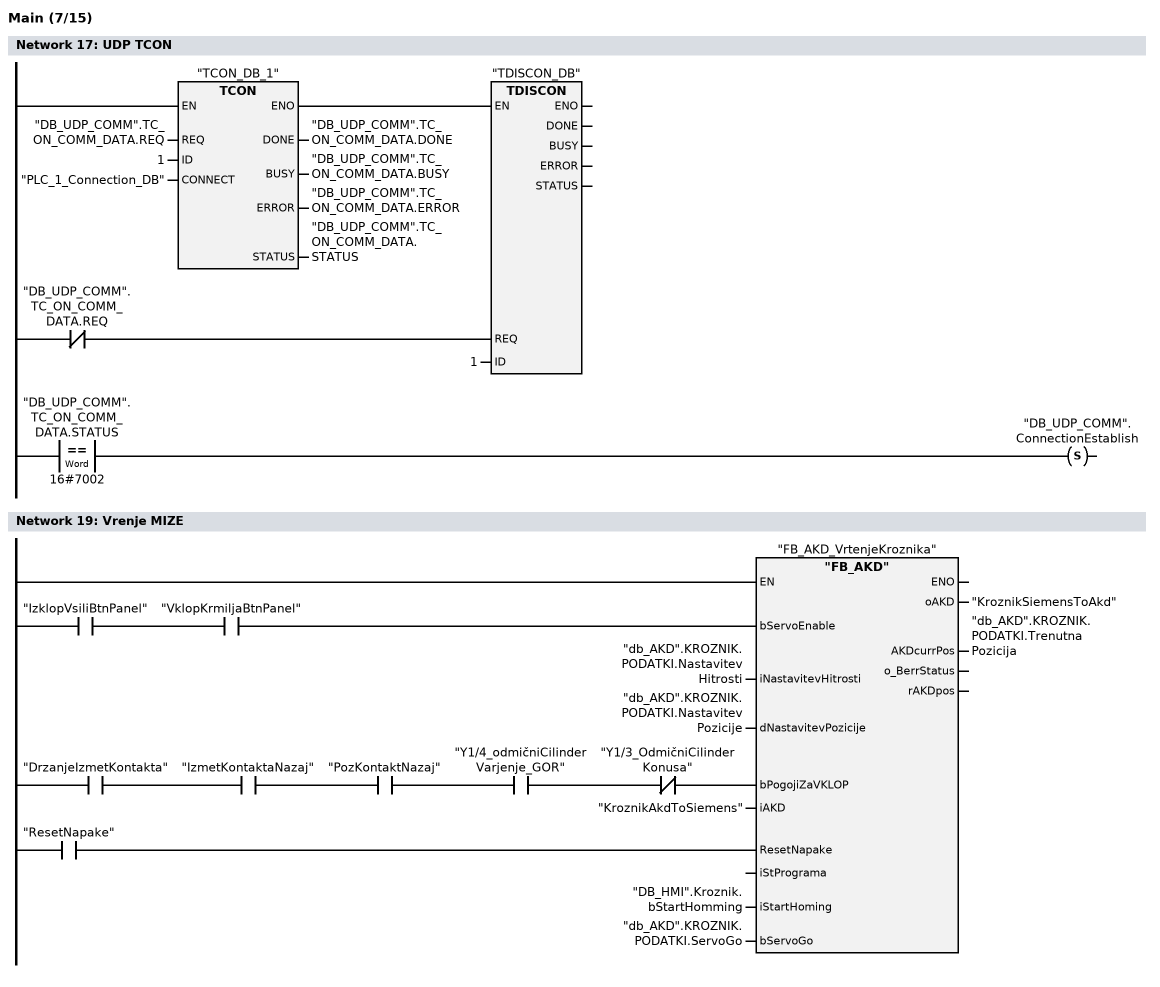
   // ENO of a box is taken as its EN; it also drops when the box reports an error
   "TCON_DB_1"(REQ := "DB_UDP_COMM".TC_ON_COMM_DATA.REQ,   // TCON
               ID := 1,
               CONNECT := "PLC_1_Connection_DB",
               DONE => "DB_UDP_COMM".TC_ON_COMM_DATA.DONE,
               BUSY => "DB_UDP_COMM".TC_ON_COMM_DATA.BUSY,
               ERROR => "DB_UDP_COMM".TC_ON_COMM_DATA.ERROR,
               STATUS => "DB_UDP_COMM".TC_ON_COMM_DATA.STATUS);
   "TDISCON_DB"(REQ := NOT "DB_UDP_COMM".TC_ON_COMM_DATA.REQ, ID := 1);   // TDISCON
   IF "DB_UDP_COMM".TC_ON_COMM_DATA.STATUS = 16#7002 THEN "DB_UDP_COMM".ConnectionEstablish := TRUE; END_IF;
END_REGION

REGION Network 18: SERVO krožna miza
END_REGION

REGION Network 19: Vrenje MIZE
   RUNG wire#powerrail
      "FB_AKD_VrtenjeKroznika"(bServoEnable := wire#w1, bPogojiZaVKLOP := wire#w2, ResetNapake := wire#w3, iNastavitevHitrosti := "db_AKD".KROZNIK.PODATKI.NastavitevHitrosti, dNastavitevPozicije := "db_AKD".KROZNIK.PODATKI.NastavitevPozicije, iAKD := "KroznikAkdToSiemens", iStPrograma :=, iStartHoming := "DB_HMI".Kroznik.bStartHomming, bServoGo := "db_AKD".KROZNIK.PODATKI.ServoGo, oAKD => "KroznikSiemensToAkd", AKDcurrPos => "db_AKD".KROZNIK.PODATKI.TrenutnaPozicija, o_BerrStatus =>, rAKDpos =>)
   END_RUNG
   RUNG wire#powerrail
      Contact( "IzklopVsiliBtnPanel" )
      Contact( "VklopKrmiljaBtnPanel" )
   END_RUNG wire#w1
   RUNG wire#powerrail
      Contact( "DrzanjeIzmetKontakta" )
      Contact( "IzmetKontaktaNazaj" )
      Contact( "PozKontaktNazaj" )
      Contact( "Y1/4_odmičniCilinderVarjenje_GOR" )
      I_Contact( "Y1/3_OdmičniCilinderKonusa" )
   END_RUNG wire#w2
   RUNG wire#powerrail
      Contact( "ResetNapake" )
   END_RUNG wire#w3
   // the same network as SCL:
   "FB_AKD_VrtenjeKroznika"(bServoEnable := "IzklopVsiliBtnPanel" AND "VklopKrmiljaBtnPanel",   // "FB_AKD"
                           iNastavitevHitrosti := "db_AKD".KROZNIK.PODATKI.NastavitevHitrosti,
                           dNastavitevPozicije := "db_AKD".KROZNIK.PODATKI.NastavitevPozicije,
                           bPogojiZaVKLOP := "DrzanjeIzmetKontakta" AND "IzmetKontaktaNazaj" AND "PozKontaktNazaj" AND "Y1/4_odmičniCilinderVarjenje_GOR" AND NOT "Y1/3_OdmičniCilinderKonusa",
                           iAKD := "KroznikAkdToSiemens",
                           ResetNapake := "ResetNapake",
                           iStartHoming := "DB_HMI".Kroznik.bStartHomming,
                           bServoGo := "db_AKD".KROZNIK.PODATKI.ServoGo,
                           oAKD => "KroznikSiemensToAkd",
                           AKDcurrPos => "db_AKD".KROZNIK.PODATKI.TrenutnaPozicija);
END_REGION

REGION Network 20: AKD REZANJE PODAJANJE
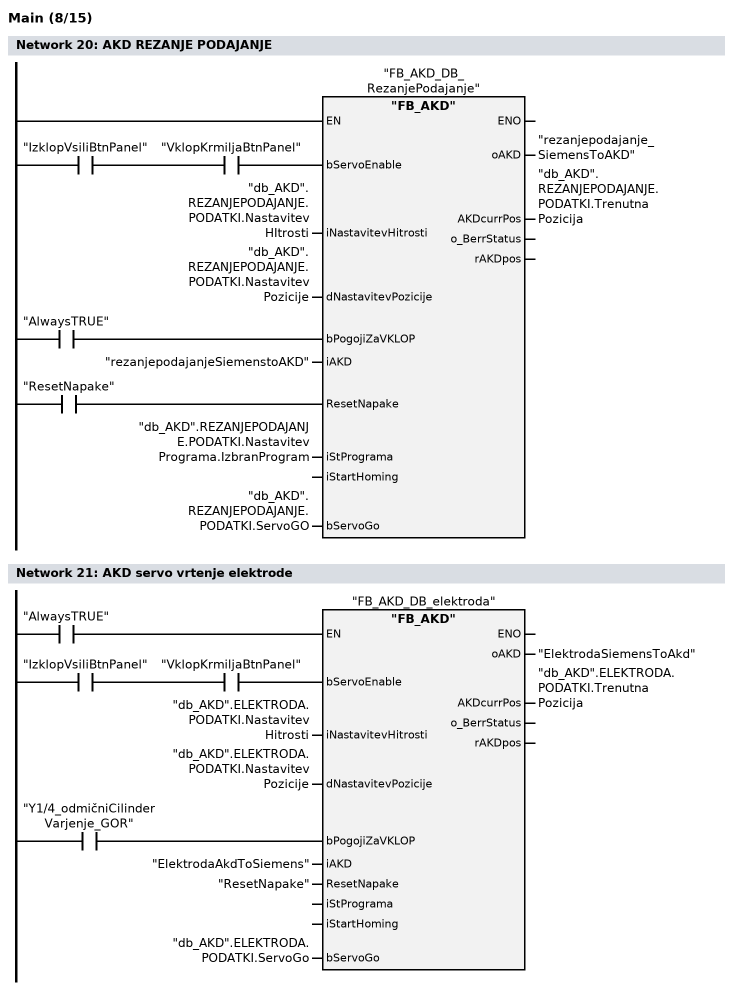
   RUNG wire#powerrail
      "FB_AKD_DB_RezanjePodajanje"(bServoEnable := wire#w1, bPogojiZaVKLOP := wire#w2, ResetNapake := wire#w3, iNastavitevHitrosti := "db_AKD".REZANJEPODAJANJE.PODATKI.NastavitevHItrosti, dNastavitevPozicije := "db_AKD".REZANJEPODAJANJE.PODATKI.NastavitevPozicije, iAKD := "rezanjepodajanjeSiemenstoAKD", iStPrograma := "db_AKD".REZANJEPODAJANJE.PODATKI.NastavitevPrograma.IzbranProgram, iStartHoming :=, bServoGo := "db_AKD".REZANJEPODAJANJE.PODATKI.ServoGO, oAKD => "rezanjepodajanje_SiemensToAKD", AKDcurrPos => "db_AKD".REZANJEPODAJANJE.PODATKI.TrenutnaPozicija, o_BerrStatus =>, rAKDpos =>)
   END_RUNG
   RUNG wire#powerrail
      Contact( "IzklopVsiliBtnPanel" )
      Contact( "VklopKrmiljaBtnPanel" )
   END_RUNG wire#w1
   RUNG wire#powerrail
      Contact( "AlwaysTRUE" )
   END_RUNG wire#w2
   RUNG wire#powerrail
      Contact( "ResetNapake" )
   END_RUNG wire#w3
   // the same network as SCL:
   "FB_AKD_DB_RezanjePodajanje"(bServoEnable := "IzklopVsiliBtnPanel" AND "VklopKrmiljaBtnPanel",   // "FB_AKD"
                           iNastavitevHitrosti := "db_AKD".REZANJEPODAJANJE.PODATKI.NastavitevHItrosti,
                           dNastavitevPozicije := "db_AKD".REZANJEPODAJANJE.PODATKI.NastavitevPozicije,
                           bPogojiZaVKLOP := "AlwaysTRUE",
                           iAKD := "rezanjepodajanjeSiemenstoAKD",
                           ResetNapake := "ResetNapake",
                           iStPrograma := "db_AKD".REZANJEPODAJANJE.PODATKI.NastavitevPrograma.IzbranProgram,
                           bServoGo := "db_AKD".REZANJEPODAJANJE.PODATKI.ServoGO,
                           oAKD => "rezanjepodajanje_SiemensToAKD",
                           AKDcurrPos => "db_AKD".REZANJEPODAJANJE.PODATKI.TrenutnaPozicija);
END_REGION

REGION Network 21: AKD servo vrtenje elektrode
   RUNG wire#powerrail
      Contact( "AlwaysTRUE" )
      "FB_AKD_DB_elektroda"(bServoEnable := wire#w1, bPogojiZaVKLOP := wire#w2, iNastavitevHitrosti := "db_AKD".ELEKTRODA.PODATKI.NastavitevHitrosti, dNastavitevPozicije := "db_AKD".ELEKTRODA.PODATKI.NastavitevPozicije, iAKD := "ElektrodaAkdToSiemens", ResetNapake := "ResetNapake", iStPrograma :=, iStartHoming :=, bServoGo := "db_AKD".ELEKTRODA.PODATKI.ServoGo, oAKD => "ElektrodaSiemensToAkd", AKDcurrPos => "db_AKD".ELEKTRODA.PODATKI.TrenutnaPozicija, o_BerrStatus =>, rAKDpos =>)
   END_RUNG
   RUNG wire#powerrail
      Contact( "IzklopVsiliBtnPanel" )
      Contact( "VklopKrmiljaBtnPanel" )
   END_RUNG wire#w1
   RUNG wire#powerrail
      Contact( "Y1/4_odmičniCilinderVarjenje_GOR" )
   END_RUNG wire#w2
   // the same network as SCL:
   IF "AlwaysTRUE" THEN
       "FB_AKD_DB_elektroda"(bServoEnable := "IzklopVsiliBtnPanel" AND "VklopKrmiljaBtnPanel",   // "FB_AKD"
                             iNastavitevHitrosti := "db_AKD".ELEKTRODA.PODATKI.NastavitevHitrosti,
                             dNastavitevPozicije := "db_AKD".ELEKTRODA.PODATKI.NastavitevPozicije,
                             bPogojiZaVKLOP := "Y1/4_odmičniCilinderVarjenje_GOR",
                             iAKD := "ElektrodaAkdToSiemens",
                             ResetNapake := "ResetNapake",
                             bServoGo := "db_AKD".ELEKTRODA.PODATKI.ServoGo,
                             oAKD => "ElektrodaSiemensToAkd",
                             AKDcurrPos => "db_AKD".ELEKTRODA.PODATKI.TrenutnaPozicija);
   END_IF;
END_REGION

REGION Network 25: SHIFT REGISTRI
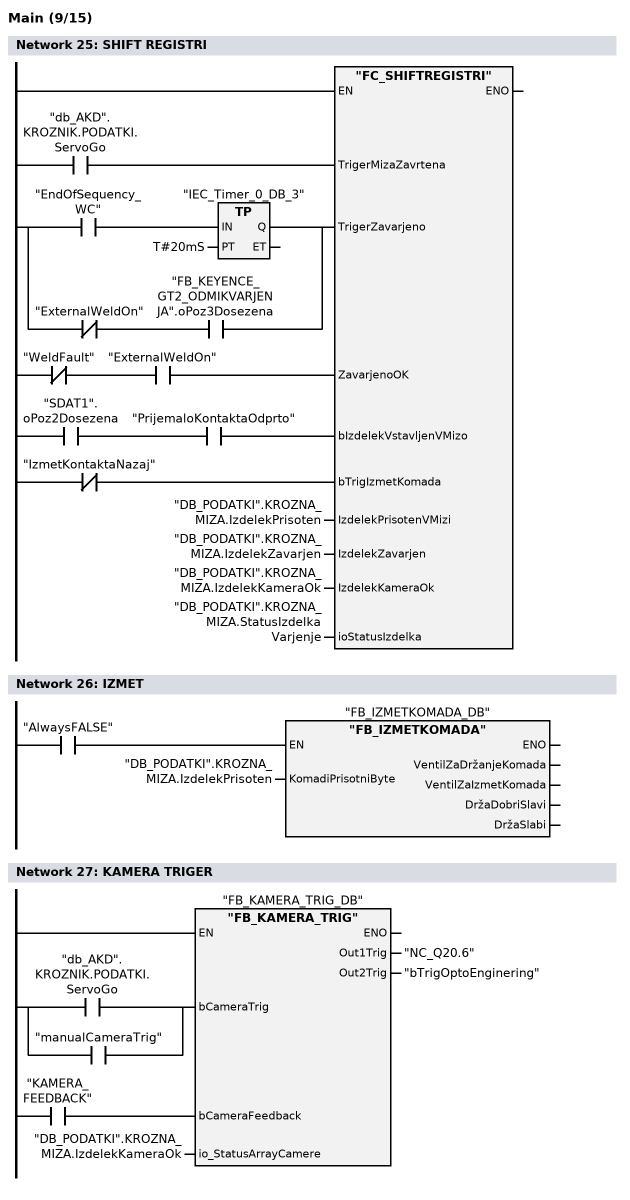
   "IEC_Timer_0_DB_3".TP(IN := "EndOfSequency_WC", PT := T#20mS);
   "FC_SHIFTREGISTRI"(TrigerMizaZavrtena := "db_AKD".KROZNIK.PODATKI.ServoGo,
                      TrigerZavarjeno := "IEC_Timer_0_DB_3".Q OR (NOT "ExternalWeldOn" AND "FB_KEYENCE_GT2_ODMIKVARJENJA".oPoz3Dosezena),
                      ZavarjenoOK := NOT "WeldFault" AND "ExternalWeldOn",
                      bIzdelekVstavljenVMizo := "SDAT1".oPoz2Dosezena AND "PrijemaloKontaktaOdprto",
                      bTrigIzmetKomada := NOT "IzmetKontaktaNazaj",
                      IzdelekPrisotenVMizi := "DB_PODATKI".KROZNA_MIZA.IzdelekPrisoten,
                      IzdelekZavarjen := "DB_PODATKI".KROZNA_MIZA.IzdelekZavarjen,
                      IzdelekKameraOk := "DB_PODATKI".KROZNA_MIZA.IzdelekKameraOk,
                      ioStatusIzdelka := "DB_PODATKI".KROZNA_MIZA.StatusIzdelkaVarjenje);
END_REGION

REGION Network 26: IZMET
   RUNG wire#powerrail
      Contact( "AlwaysFALSE" )
      "FB_IZMETKOMADA_DB"(KomadiPrisotniByte := "DB_PODATKI".KROZNA_MIZA.IzdelekPrisoten, VentilZaDržanjeKomada =>, VentilZaIzmetKomada =>, DržaDobriSlavi =>, DržaSlabi =>)
   END_RUNG
   // the same network as SCL:
   IF "AlwaysFALSE" THEN
       "FB_IZMETKOMADA_DB"(KomadiPrisotniByte := "DB_PODATKI".KROZNA_MIZA.IzdelekPrisoten);   // "FB_IZMETKOMADA"
   END_IF;
END_REGION

REGION Network 27: KAMERA TRIGER
   RUNG wire#powerrail
      "FB_KAMERA_TRIG_DB"(bCameraTrig := wire#w1, bCameraFeedback := wire#w2, io_StatusArrayCamere := "DB_PODATKI".KROZNA_MIZA.IzdelekKameraOk, Out1Trig => "NC_Q20.6", Out2Trig => "bTrigOptoEnginering")
   END_RUNG
   RUNG wire#powerrail
      Contact( "db_AKD".KROZNIK.PODATKI.ServoGo )
   END_RUNG wire#w1
   RUNG wire#powerrail
      Contact( "manualCameraTrig" )
   END_RUNG wire#w1
   RUNG wire#powerrail
      Contact( "KAMERA_FEEDBACK" )
   END_RUNG wire#w2
   // the same network as SCL:
   "FB_KAMERA_TRIG_DB"(bCameraTrig := "db_AKD".KROZNIK.PODATKI.ServoGo OR "manualCameraTrig",   // "FB_KAMERA_TRIG"
                       bCameraFeedback := "KAMERA_FEEDBACK",
                       io_StatusArrayCamere := "DB_PODATKI".KROZNA_MIZA.IzdelekKameraOk,
                       Out1Trig => "NC_Q20.6",
                       Out2Trig => "bTrigOptoEnginering");
END_REGION

REGION Network 31: AKD - podajanjerezanje
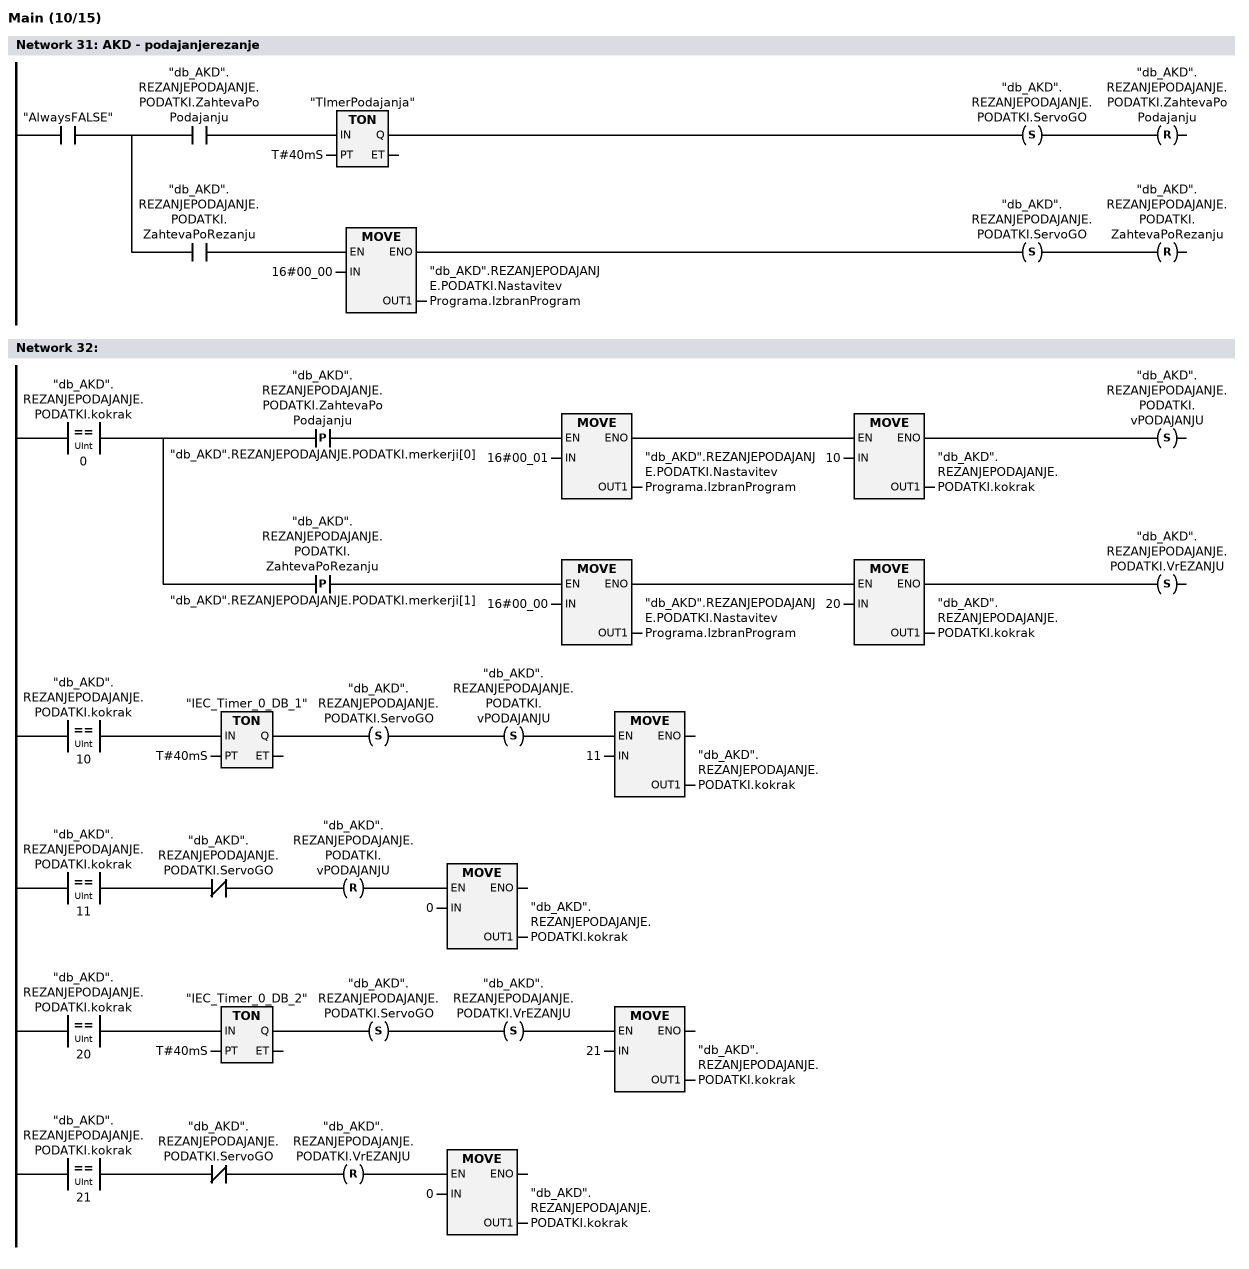
   "TImerPodajanja".TON(IN := "AlwaysFALSE" AND "db_AKD".REZANJEPODAJANJE.PODATKI.ZahtevaPoPodajanju,
                        PT := T#40mS);
   IF "TImerPodajanja".Q THEN
       "db_AKD".REZANJEPODAJANJE.PODATKI.ServoGO := TRUE;
       "db_AKD".REZANJEPODAJANJE.PODATKI.ZahtevaPoPodajanju := FALSE;
   END_IF;
   IF "AlwaysFALSE" AND "db_AKD".REZANJEPODAJANJE.PODATKI.ZahtevaPoRezanju THEN
       "db_AKD".REZANJEPODAJANJE.PODATKI.NastavitevPrograma.IzbranProgram := 16#00_00;
       "db_AKD".REZANJEPODAJANJE.PODATKI.ServoGO := TRUE;
       "db_AKD".REZANJEPODAJANJE.PODATKI.ZahtevaPoRezanju := FALSE;
   END_IF;
END_REGION

REGION Network 32
   #_w1 := "db_AKD".REZANJEPODAJANJE.PODATKI.kokrak = 0;
   #_w2 := #_w1 AND "db_AKD".REZANJEPODAJANJE.PODATKI.ZahtevaPoPodajanju AND NOT "db_AKD".REZANJEPODAJANJE.PODATKI.merkerji[0];   // rising edge of "db_AKD".REZANJEPODAJANJE.PODATKI.ZahtevaPoPodajanju
   "db_AKD".REZANJEPODAJANJE.PODATKI.merkerji[0] := "db_AKD".REZANJEPODAJANJE.PODATKI.ZahtevaPoPodajanju;
   IF #_w2 THEN
       "db_AKD".REZANJEPODAJANJE.PODATKI.NastavitevPrograma.IzbranProgram := 16#00_01;
       "db_AKD".REZANJEPODAJANJE.PODATKI.kokrak := 10;
       "db_AKD".REZANJEPODAJANJE.PODATKI.vPODAJANJU := TRUE;
   END_IF;
   #_w3 := #_w1 AND "db_AKD".REZANJEPODAJANJE.PODATKI.ZahtevaPoRezanju AND NOT "db_AKD".REZANJEPODAJANJE.PODATKI.merkerji[1];   // rising edge of "db_AKD".REZANJEPODAJANJE.PODATKI.ZahtevaPoRezanju
   "db_AKD".REZANJEPODAJANJE.PODATKI.merkerji[1] := "db_AKD".REZANJEPODAJANJE.PODATKI.ZahtevaPoRezanju;
   IF #_w3 THEN
       "db_AKD".REZANJEPODAJANJE.PODATKI.NastavitevPrograma.IzbranProgram := 16#00_00;
       "db_AKD".REZANJEPODAJANJE.PODATKI.kokrak := 20;
       "db_AKD".REZANJEPODAJANJE.PODATKI.VrEZANJU := TRUE;
   END_IF;
   "IEC_Timer_0_DB_1".TON(IN := "db_AKD".REZANJEPODAJANJE.PODATKI.kokrak = 10, PT := T#40mS);
   IF "IEC_Timer_0_DB_1".Q THEN
       "db_AKD".REZANJEPODAJANJE.PODATKI.ServoGO := TRUE;
       "db_AKD".REZANJEPODAJANJE.PODATKI.vPODAJANJU := TRUE;
       "db_AKD".REZANJEPODAJANJE.PODATKI.kokrak := 11;
   END_IF;
   IF ("db_AKD".REZANJEPODAJANJE.PODATKI.kokrak = 11) AND NOT "db_AKD".REZANJEPODAJANJE.PODATKI.ServoGO THEN
       "db_AKD".REZANJEPODAJANJE.PODATKI.vPODAJANJU := FALSE;
       "db_AKD".REZANJEPODAJANJE.PODATKI.kokrak := 0;
   END_IF;
   "IEC_Timer_0_DB_2".TON(IN := "db_AKD".REZANJEPODAJANJE.PODATKI.kokrak = 20, PT := T#40mS);
   IF "IEC_Timer_0_DB_2".Q THEN
       "db_AKD".REZANJEPODAJANJE.PODATKI.ServoGO := TRUE;
       "db_AKD".REZANJEPODAJANJE.PODATKI.VrEZANJU := TRUE;
       "db_AKD".REZANJEPODAJANJE.PODATKI.kokrak := 21;
   END_IF;
   IF ("db_AKD".REZANJEPODAJANJE.PODATKI.kokrak = 21) AND NOT "db_AKD".REZANJEPODAJANJE.PODATKI.ServoGO THEN
       "db_AKD".REZANJEPODAJANJE.PODATKI.VrEZANJU := FALSE;
       "db_AKD".REZANJEPODAJANJE.PODATKI.kokrak := 0;
   END_IF;
END_REGION

REGION Network 33 (SCL): REZANJE/PODAJANJE
END_REGION

REGION Network 34: VARJENJE - bosh
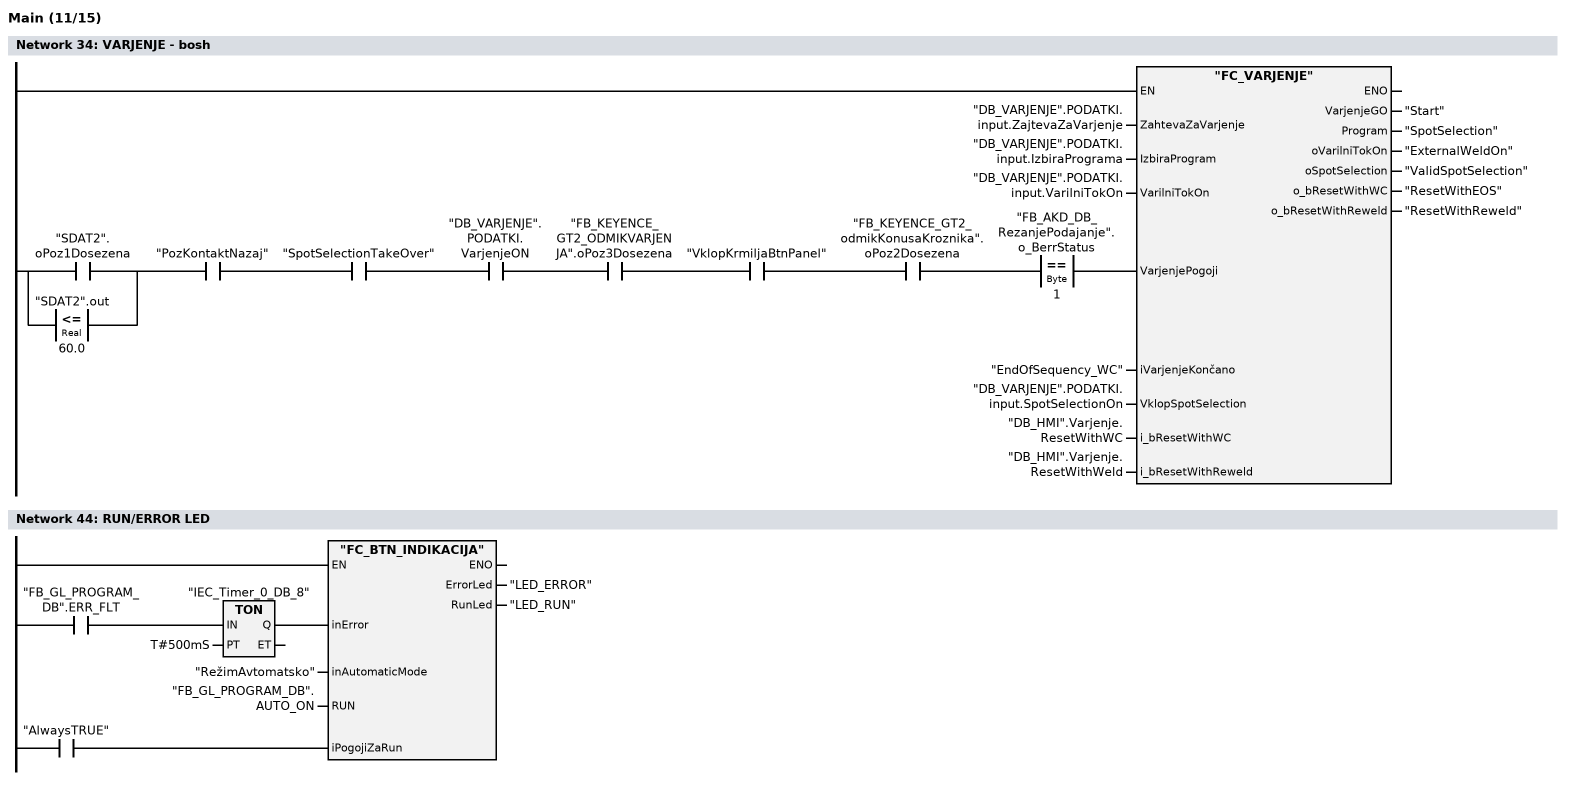
   RUNG wire#powerrail
      "FC_VARJENJE"(VarjenjePogoji := wire#w2, ZahtevaZaVarjenje := "DB_VARJENJE".PODATKI.input.ZajtevaZaVarjenje, IzbiraProgram := "DB_VARJENJE".PODATKI.input.IzbiraPrograma, VarilniTokOn := "DB_VARJENJE".PODATKI.input.VarilniTokOn, iVarjenjeKončano := "EndOfSequency_WC", VklopSpotSelection := "DB_VARJENJE".PODATKI.input.SpotSelectionOn, i_bResetWithWC := "DB_HMI".Varjenje.ResetWithWC, i_bResetWithReweld := "DB_HMI".Varjenje.ResetWithWeld, VarjenjeGO => "Start", Program => "SpotSelection", oVarilniTokOn => "ExternalWeldOn", oSpotSelection => "ValidSpotSelection", o_bResetWithWC => "ResetWithEOS", o_bResetWithReweld => "ResetWithReweld")
   END_RUNG
   RUNG wire#powerrail
      Contact( "SDAT2".oPoz1Dosezena )
      wire#w1
      Contact( "PozKontaktNazaj" )
      Contact( "SpotSelectionTakeOver" )
      Contact( "DB_VARJENJE".PODATKI.VarjenjeON )
      Contact( "FB_KEYENCE_GT2_ODMIKVARJENJA".oPoz3Dosezena )
      Contact( "VklopKrmiljaBtnPanel" )
      Contact( "FB_KEYENCE_GT2_odmikKonusaKroznika".oPoz2Dosezena )
      { S7_Templates := "SrcType := Byte" } EQ_Contact(in1 := "FB_AKD_DB_RezanjePodajanje".o_BerrStatus, in2 := 1)
   END_RUNG wire#w2
   RUNG wire#powerrail
      { S7_Templates := "SrcType := Real" } LE_Contact(in1 := "SDAT2".out, in2 := 60.0)
   END_RUNG wire#w1
   // the same network as SCL:
   "FC_VARJENJE"(ZahtevaZaVarjenje := "DB_VARJENJE".PODATKI.input.ZajtevaZaVarjenje,
                 IzbiraProgram := "DB_VARJENJE".PODATKI.input.IzbiraPrograma,
                 VarilniTokOn := "DB_VARJENJE".PODATKI.input.VarilniTokOn,
                 VarjenjePogoji := ("SDAT2".oPoz1Dosezena OR ("SDAT2".out <= 60.0)) AND "PozKontaktNazaj" AND "SpotSelectionTakeOver" AND "DB_VARJENJE".PODATKI.VarjenjeON AND "FB_KEYENCE_GT2_ODMIKVARJENJA".oPoz3Dosezena AND "VklopKrmiljaBtnPanel" AND "FB_KEYENCE_GT2_odmikKonusaKroznika".oPoz2Dosezena AND ("FB_AKD_DB_RezanjePodajanje".o_BerrStatus = 1),
                 iVarjenjeKončano := "EndOfSequency_WC",
                 VklopSpotSelection := "DB_VARJENJE".PODATKI.input.SpotSelectionOn,
                 i_bResetWithWC := "DB_HMI".Varjenje.ResetWithWC,
                 i_bResetWithReweld := "DB_HMI".Varjenje.ResetWithWeld,
                 VarjenjeGO => "Start",
                 Program => "SpotSelection",
                 oVarilniTokOn => "ExternalWeldOn",
                 oSpotSelection => "ValidSpotSelection",
                 o_bResetWithWC => "ResetWithEOS",
                 o_bResetWithReweld => "ResetWithReweld");
END_REGION

REGION Network 44: RUN/ERROR LED
   "IEC_Timer_0_DB_8".TON(IN := "FB_GL_PROGRAM_DB".ERR_FLT, PT := T#500mS);
   "FC_BTN_INDIKACIJA"(inError := "IEC_Timer_0_DB_8".Q,
                       inAutomaticMode := "RežimAvtomatsko",
                       RUN := "FB_GL_PROGRAM_DB".AUTO_ON,
                       iPogojiZaRun := "AlwaysTRUE",
                       ErrorLed => "LED_ERROR",
                       RunLed => "LED_RUN");
END_REGION

REGION Network 45: IOL_BANNER
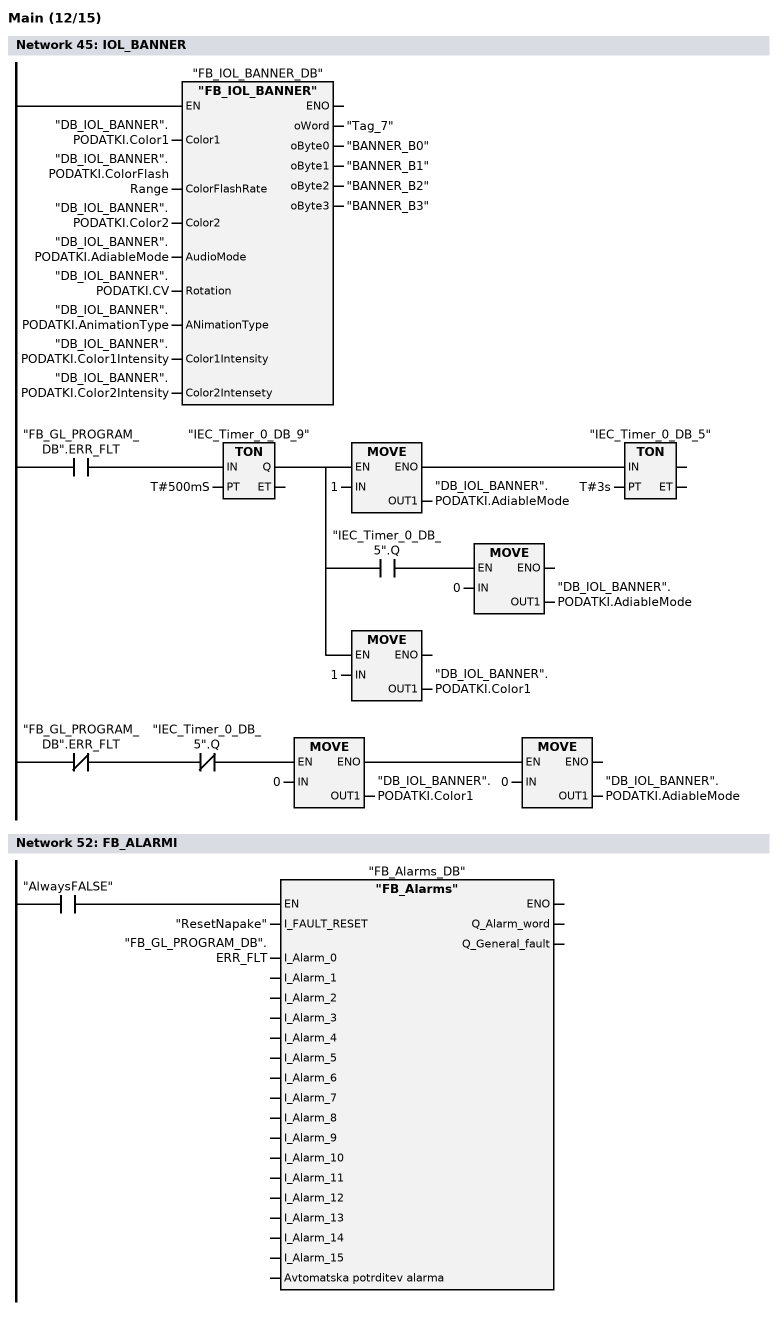
   "FB_IOL_BANNER_DB"(Color1 := "DB_IOL_BANNER".PODATKI.Color1,   // "FB_IOL_BANNER"
                      ColorFlashRate := "DB_IOL_BANNER".PODATKI.ColorFlashRange,
                      Color2 := "DB_IOL_BANNER".PODATKI.Color2,
                      AudioMode := "DB_IOL_BANNER".PODATKI.AdiableMode,
                      Rotation := "DB_IOL_BANNER".PODATKI.CV,
                      ANimationType := "DB_IOL_BANNER".PODATKI.AnimationType,
                      Color1Intensity := "DB_IOL_BANNER".PODATKI.Color1Intensity,
                      Color2Intensety := "DB_IOL_BANNER".PODATKI.Color2Intensity,
                      oWord => "Tag_7",
                      oByte0 => "BANNER_B0",
                      oByte1 => "BANNER_B1",
                      oByte2 => "BANNER_B2",
                      oByte3 => "BANNER_B3");
   "IEC_Timer_0_DB_9".TON(IN := "FB_GL_PROGRAM_DB".ERR_FLT, PT := T#500mS);
   IF "IEC_Timer_0_DB_9".Q THEN "DB_IOL_BANNER".PODATKI.AdiableMode := 1; END_IF;
   "IEC_Timer_0_DB_5".TON(IN := "IEC_Timer_0_DB_9".Q, PT := T#3s);
   IF "IEC_Timer_0_DB_9".Q AND "IEC_Timer_0_DB_5".Q THEN "DB_IOL_BANNER".PODATKI.AdiableMode := 0; END_IF;
   IF "IEC_Timer_0_DB_9".Q THEN "DB_IOL_BANNER".PODATKI.Color1 := 1; END_IF;
   IF NOT "FB_GL_PROGRAM_DB".ERR_FLT AND NOT "IEC_Timer_0_DB_5".Q THEN
       "DB_IOL_BANNER".PODATKI.Color1 := 0;
       "DB_IOL_BANNER".PODATKI.AdiableMode := 0;
   END_IF;
END_REGION

REGION Network 51: FB_ALARMI
END_REGION

REGION Network 52: FB_ALARMI
   RUNG wire#powerrail
      Contact( "AlwaysFALSE" )
      "FB_Alarms_DB"(I_FAULT_RESET := "ResetNapake", I_Alarm_0 := "FB_GL_PROGRAM_DB".ERR_FLT, I_Alarm_1 :=, I_Alarm_2 :=, I_Alarm_3 :=, I_Alarm_4 :=, I_Alarm_5 :=, I_Alarm_6 :=, I_Alarm_7 :=, I_Alarm_8 :=, I_Alarm_9 :=, I_Alarm_10 :=, I_Alarm_11 :=, I_Alarm_12 :=, I_Alarm_13 :=, I_Alarm_14 :=, I_Alarm_15 :=, "Avtomatska potrditev alarma" :=, Q_Alarm_word =>, Q_General_fault =>)
   END_RUNG
   // the same network as SCL:
   IF "AlwaysFALSE" THEN
       "FB_Alarms_DB"(I_FAULT_RESET := "ResetNapake", I_Alarm_0 := "FB_GL_PROGRAM_DB".ERR_FLT);   // "FB_Alarms"
   END_IF;
END_REGION

REGION Network 55: HOMING - RESETIRANJE VREDNOSTI V MIZI
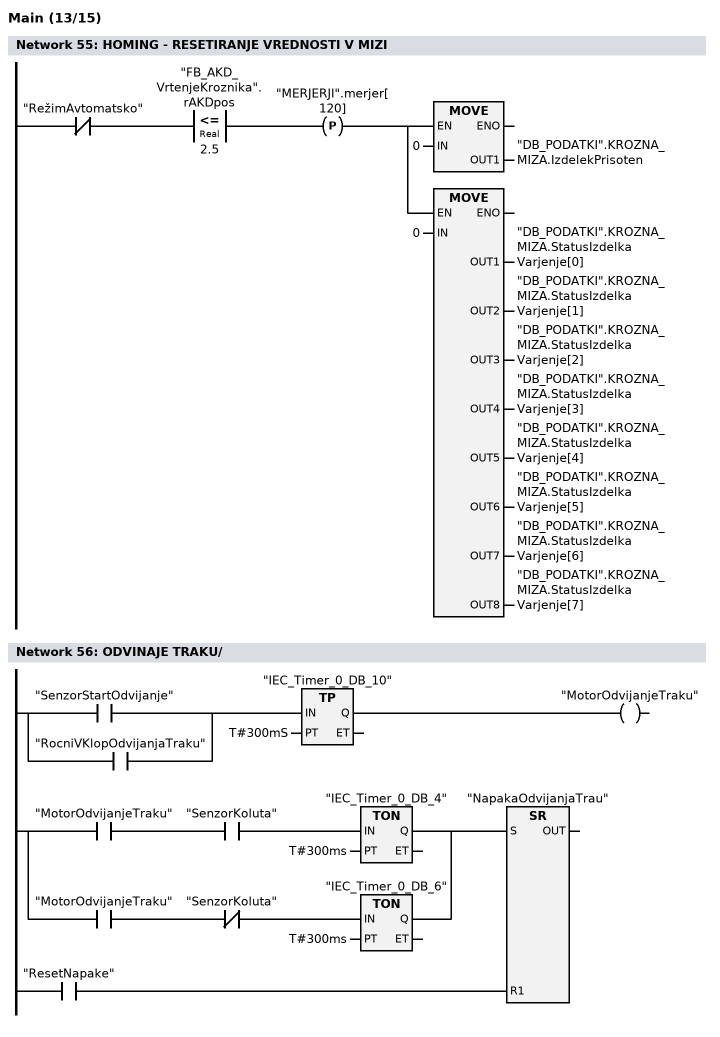
   RUNG wire#powerrail
      I_Contact( "RežimAvtomatsko" )
      { S7_Templates := "SrcType := Real" } LE_Contact(in1 := "FB_AKD_VrtenjeKroznika".rAKDpos, in2 := 2.5)
      P_Trig( "MERJERJI".merjer[120] )
      wire#w1
      Move(in := 0, out1 => "DB_PODATKI".KROZNA_MIZA.IzdelekPrisoten)
   END_RUNG
   RUNG wire#w1
      Move(in := 0, out1 => "DB_PODATKI".KROZNA_MIZA.StatusIzdelkaVarjenje[0], out2 => "DB_PODATKI".KROZNA_MIZA.StatusIzdelkaVarjenje[1], out3 => "DB_PODATKI".KROZNA_MIZA.StatusIzdelkaVarjenje[2], out4 => "DB_PODATKI".KROZNA_MIZA.StatusIzdelkaVarjenje[3], out5 => "DB_PODATKI".KROZNA_MIZA.StatusIzdelkaVarjenje[4], out6 => "DB_PODATKI".KROZNA_MIZA.StatusIzdelkaVarjenje[5], out7 => "DB_PODATKI".KROZNA_MIZA.StatusIzdelkaVarjenje[6], out8 => "DB_PODATKI".KROZNA_MIZA.StatusIzdelkaVarjenje[7])
   END_RUNG
   // the same network as SCL:
   #_w1 := NOT "RežimAvtomatsko" AND ("FB_AKD_VrtenjeKroznika".rAKDpos <= 2.5);
   #_w2 := #_w1 AND NOT "MERJERJI".merjer[120];   // rising edge
   "MERJERJI".merjer[120] := #_w1;
   IF #_w2 THEN
       "DB_PODATKI".KROZNA_MIZA.IzdelekPrisoten := 0;
       "DB_PODATKI".KROZNA_MIZA.StatusIzdelkaVarjenje[0] := 0;
       "DB_PODATKI".KROZNA_MIZA.StatusIzdelkaVarjenje[1] := 0;
       "DB_PODATKI".KROZNA_MIZA.StatusIzdelkaVarjenje[2] := 0;
       "DB_PODATKI".KROZNA_MIZA.StatusIzdelkaVarjenje[3] := 0;
       "DB_PODATKI".KROZNA_MIZA.StatusIzdelkaVarjenje[4] := 0;
       "DB_PODATKI".KROZNA_MIZA.StatusIzdelkaVarjenje[5] := 0;
       "DB_PODATKI".KROZNA_MIZA.StatusIzdelkaVarjenje[6] := 0;
       "DB_PODATKI".KROZNA_MIZA.StatusIzdelkaVarjenje[7] := 0;
   END_IF;
END_REGION

REGION Network 56: ODVINAJE TRAKU/
   "IEC_Timer_0_DB_10".TP(IN := "SenzorStartOdvijanje" OR "RocniVKlopOdvijanjaTraku", PT := T#300mS);
   "MotorOdvijanjeTraku" := "IEC_Timer_0_DB_10".Q;
   "IEC_Timer_0_DB_4".TON(IN := "MotorOdvijanjeTraku" AND "SenzorKoluta", PT := T#300ms);
   "IEC_Timer_0_DB_6".TON(IN := "MotorOdvijanjeTraku" AND NOT "SenzorKoluta", PT := T#300ms);
   IF "IEC_Timer_0_DB_4".Q OR "IEC_Timer_0_DB_6".Q THEN
       "NapakaOdvijanjaTrau" := TRUE;   // SR flip-flop
   END_IF;
   IF "ResetNapake" THEN "NapakaOdvijanjaTrau" := FALSE; END_IF;
END_REGION

REGION Network 57: Odvijanje Čiščenje Elektrode